REGION Network 31: Positioning commands
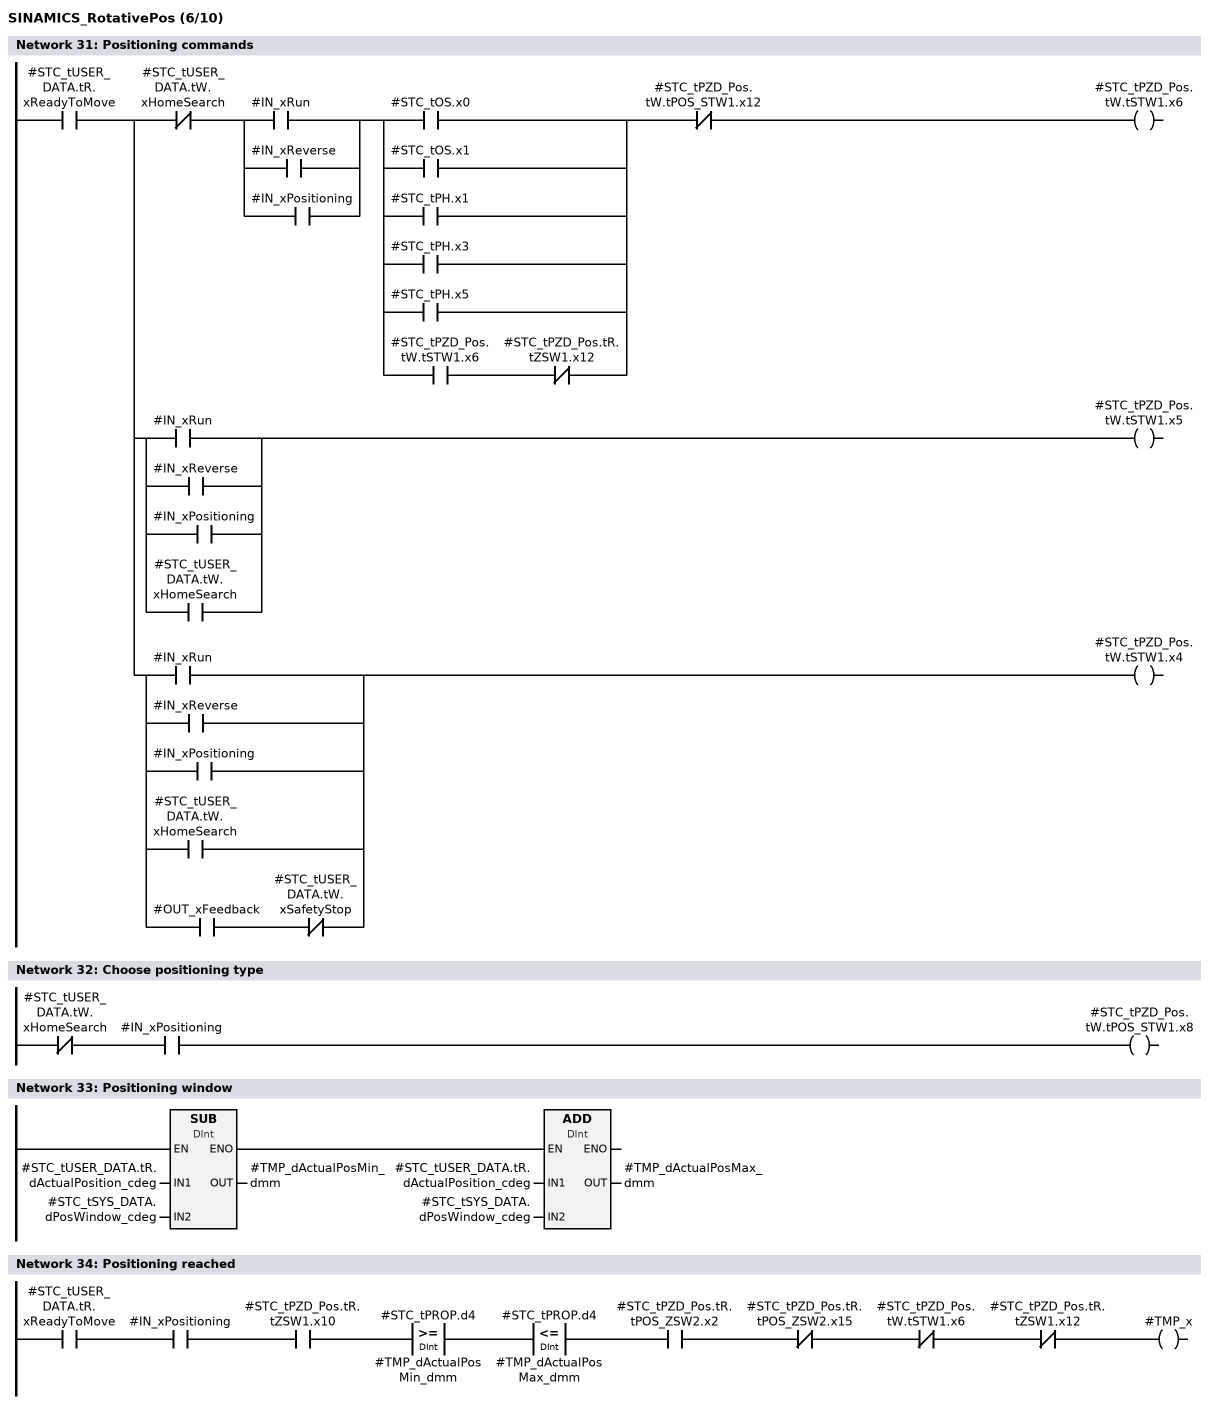
   RUNG wire#powerrail
      Contact( #STC_tUSER_DATA.tR.xReadyToMove )
      wire#w1
      I_Contact( #STC_tUSER_DATA.tW.xHomeSearch )
      wire#w2
      Contact( #IN_xRun )
      wire#w3
      Contact( #STC_tOS.x0 )
      wire#w4
      I_Contact( #STC_tPZD_Pos.tW.tPOS_STW1.x12 )
      Coil( #STC_tPZD_Pos.tW.tSTW1.x6 )
   END_RUNG
   RUNG wire#w2
      Contact( #IN_xReverse )
   END_RUNG wire#w3
   RUNG wire#w2
      Contact( #IN_xPositioning )
   END_RUNG wire#w3
   RUNG wire#w3
      Contact( #STC_tOS.x1 )
   END_RUNG wire#w4
   RUNG wire#w3
      Contact( #STC_tPH.x1 )
   END_RUNG wire#w4
   RUNG wire#w3
      Contact( #STC_tPH.x3 )
   END_RUNG wire#w4
   RUNG wire#w3
      Contact( #STC_tPH.x5 )
   END_RUNG wire#w4
   RUNG wire#w3
      Contact( #STC_tPZD_Pos.tW.tSTW1.x6 )
      I_Contact( #STC_tPZD_Pos.tR.tZSW1.x12 )
   END_RUNG wire#w4
   RUNG wire#w1
      Contact( #IN_xRun )
      wire#w5
      Coil( #STC_tPZD_Pos.tW.tSTW1.x5 )
   END_RUNG
   RUNG wire#w1
      Contact( #IN_xReverse )
   END_RUNG wire#w5
   RUNG wire#w1
      Contact( #IN_xPositioning )
   END_RUNG wire#w5
   RUNG wire#w1
      Contact( #STC_tUSER_DATA.tW.xHomeSearch )
   END_RUNG wire#w5
   RUNG wire#w1
      Contact( #IN_xRun )
      wire#w6
      Coil( #STC_tPZD_Pos.tW.tSTW1.x4 )
   END_RUNG
   RUNG wire#w1
      Contact( #IN_xReverse )
   END_RUNG wire#w6
   RUNG wire#w1
      Contact( #IN_xPositioning )
   END_RUNG wire#w6
   RUNG wire#w1
      Contact( #STC_tUSER_DATA.tW.xHomeSearch )
   END_RUNG wire#w6
   RUNG wire#w1
      Contact( #OUT_xFeedback )
      I_Contact( #STC_tUSER_DATA.tW.xSafetyStop )
   END_RUNG wire#w6
   // the same network as SCL:
   #STC_tPZD_Pos.tW.tSTW1.x6 := #STC_tUSER_DATA.tR.xReadyToMove AND NOT #STC_tUSER_DATA.tW.xHomeSearch AND (#IN_xRun OR #IN_xReverse OR #IN_xPositioning) AND (#STC_tOS.x0 OR #STC_tOS.x1 OR #STC_tPH.x1 OR #STC_tPH.x3 OR #STC_tPH.x5 OR (#STC_tPZD_Pos.tW.tSTW1.x6 AND NOT #STC_tPZD_Pos.tR.tZSW1.x12)) AND NOT #STC_tPZD_Pos.tW.tPOS_STW1.x12;
   #STC_tPZD_Pos.tW.tSTW1.x5 := #STC_tUSER_DATA.tR.xReadyToMove AND (#IN_xRun OR #IN_xReverse OR #IN_xPositioning OR #STC_tUSER_DATA.tW.xHomeSearch);
   #STC_tPZD_Pos.tW.tSTW1.x4 := #STC_tUSER_DATA.tR.xReadyToMove AND (#IN_xRun OR #IN_xReverse OR #IN_xPositioning OR #STC_tUSER_DATA.tW.xHomeSearch OR (#OUT_xFeedback AND NOT #STC_tUSER_DATA.tW.xSafetyStop));
END_REGION

REGION Network 32: Choose positioning type
   RUNG wire#powerrail
      I_Contact( #STC_tUSER_DATA.tW.xHomeSearch )
      Contact( #IN_xPositioning )
      Coil( #STC_tPZD_Pos.tW.tPOS_STW1.x8 )
   END_RUNG
   // the same network as SCL:
   #STC_tPZD_Pos.tW.tPOS_STW1.x8 := NOT #STC_tUSER_DATA.tW.xHomeSearch AND #IN_xPositioning;
END_REGION

REGION Network 33: Positioning window
   RUNG wire#powerrail
      { S7_Templates := "SrcType := DInt"; S7_GenerateENO := "TRUE" } Sub(in1 := #STC_tUSER_DATA.tR.dActualPosition_cdeg, in2 := #STC_tSYS_DATA.dPosWindow_cdeg, out => #TMP_dActualPosMin_dmm)
      { S7_Templates := "SrcType := DInt"; S7_GenerateENO := "TRUE" } Add(in1 := #STC_tUSER_DATA.tR.dActualPosition_cdeg, in2 := #STC_tSYS_DATA.dPosWindow_cdeg, out => #TMP_dActualPosMax_dmm)
   END_RUNG
   // the same network as SCL:
   // ENO of a box is taken as its EN; it also drops when the box reports an error
   #TMP_dActualPosMin_dmm := #STC_tUSER_DATA.tR.dActualPosition_cdeg - #STC_tSYS_DATA.dPosWindow_cdeg;
   #TMP_dActualPosMax_dmm := #STC_tUSER_DATA.tR.dActualPosition_cdeg + #STC_tSYS_DATA.dPosWindow_cdeg;
END_REGION

REGION Network 34: Positioning reached
   RUNG wire#powerrail
      Contact( #STC_tUSER_DATA.tR.xReadyToMove )
      Contact( #IN_xPositioning )
      Contact( #STC_tPZD_Pos.tR.tZSW1.x10 )
      { S7_Templates := "SrcType := DInt" } GE_Contact(in1 := #STC_tPROP.d4, in2 := #TMP_dActualPosMin_dmm)
      { S7_Templates := "SrcType := DInt" } LE_Contact(in1 := #STC_tPROP.d4, in2 := #TMP_dActualPosMax_dmm)
      Contact( #STC_tPZD_Pos.tR.tPOS_ZSW2.x2 )
      I_Contact( #STC_tPZD_Pos.tR.tPOS_ZSW2.x15 )
      I_Contact( #STC_tPZD_Pos.tW.tSTW1.x6 )
      I_Contact( #STC_tPZD_Pos.tR.tZSW1.x12 )
      Coil( #TMP_x )
   END_RUNG
   // the same network as SCL:
   #TMP_x := #STC_tUSER_DATA.tR.xReadyToMove AND #IN_xPositioning AND #STC_tPZD_Pos.tR.tZSW1.x10 AND (#STC_tPROP.d4 >= #TMP_dActualPosMin_dmm) AND (#STC_tPROP.d4 <= #TMP_dActualPosMax_dmm) AND #STC_tPZD_Pos.tR.tPOS_ZSW2.x2 AND NOT #STC_tPZD_Pos.tR.tPOS_ZSW2.x15 AND NOT #STC_tPZD_Pos.tW.tSTW1.x6 AND NOT #STC_tPZD_Pos.tR.tZSW1.x12;
END_REGION

REGION Network 35: Positioning reached
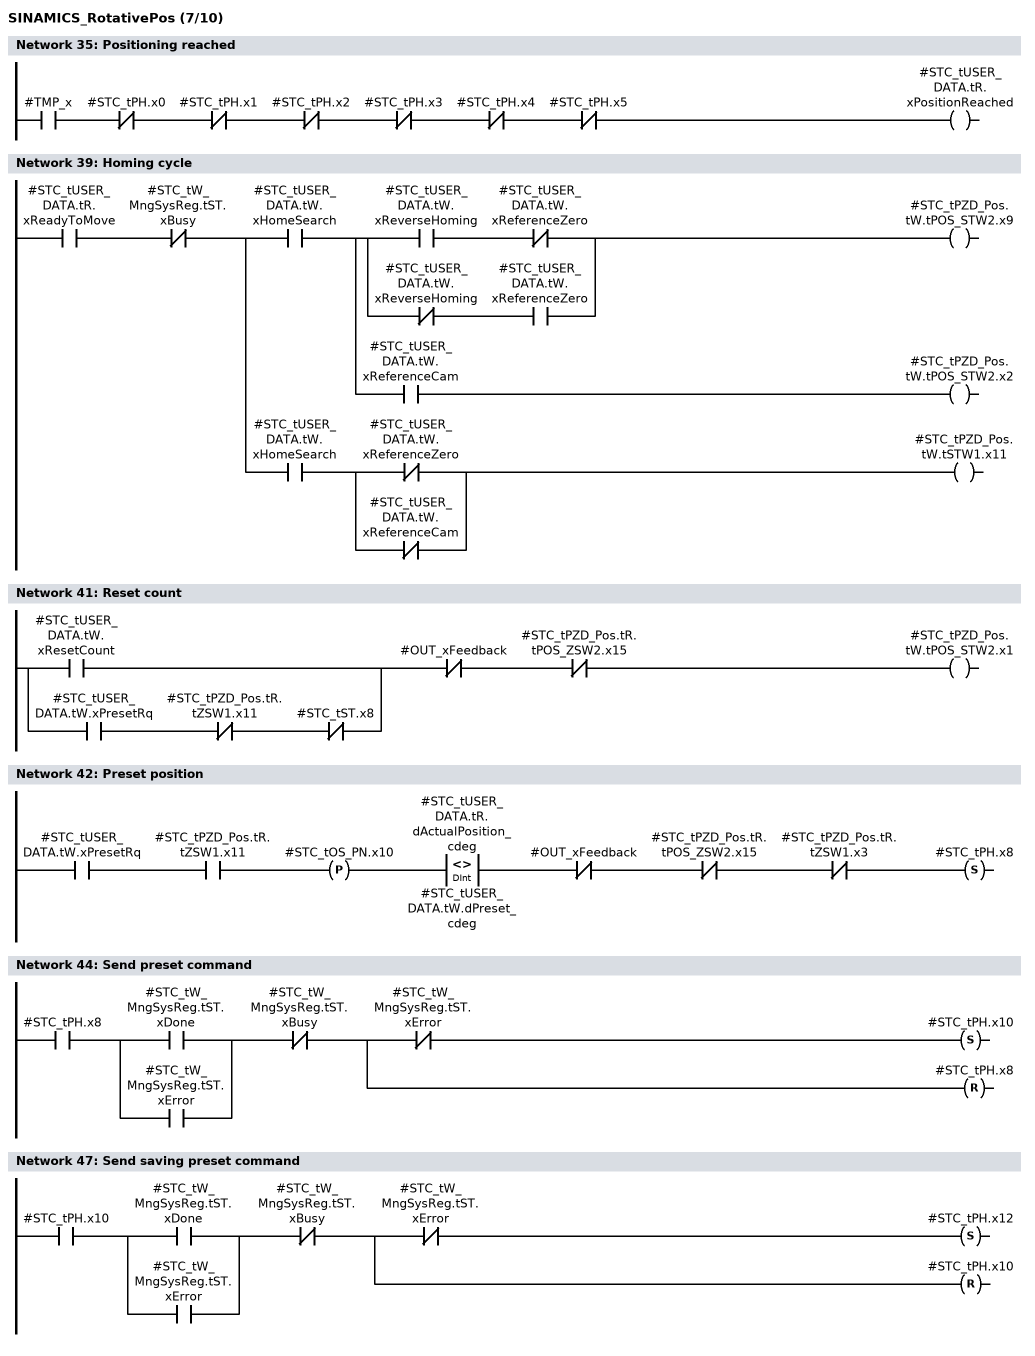
   RUNG wire#powerrail
      Contact( #TMP_x )
      I_Contact( #STC_tPH.x0 )
      I_Contact( #STC_tPH.x1 )
      I_Contact( #STC_tPH.x2 )
      I_Contact( #STC_tPH.x3 )
      I_Contact( #STC_tPH.x4 )
      I_Contact( #STC_tPH.x5 )
      Coil( #STC_tUSER_DATA.tR.xPositionReached )
   END_RUNG
   // the same network as SCL:
   #STC_tUSER_DATA.tR.xPositionReached := #TMP_x AND NOT #STC_tPH.x0 AND NOT #STC_tPH.x1 AND NOT #STC_tPH.x2 AND NOT #STC_tPH.x3 AND NOT #STC_tPH.x4 AND NOT #STC_tPH.x5;
END_REGION

REGION Network 36: #####_HOMING_CYCLE_#####
END_REGION

REGION Network 37 (STL): Send homing preset
         A     #STC_tUSER_DATA.tW.xHomeSearch;
         AN    #STC_tPZD_Pos.tW.tSTW1.x11;
         JCN   PrH0;
         =     #STC_tW_MngSysReg.tST.xWrite_Request;

         L     #STC_tSYS_DATA.iPosPZD_MM;
         SLW   8;
         L     W#16#2;
         OW;
         T     #STC_tW_MngSysReg.tDATA.wRequest_refere_RequestID;
         L     #STC_tSYS_DATA.iPosPZD_MM;
         SLW   8;
         L     W#16#1;
         OW;
         T     #STC_tW_MngSysReg.tDATA.wAxis_NoOfParameters;
         L     W#16#1001;
         T     #STC_tW_MngSysReg.tDATA.wAttribute_NoOfElements;
         L     2599;
         T     #STC_tW_MngSysReg.tDATA.iParameter_number;
         L     W#16#0;
         T     #STC_tW_MngSysReg.tDATA.wSubindex;
         L     W#16#4301;
         T     #STC_tW_MngSysReg.tDATA.wFormat_NoOfValue;
         L     #STC_tSYS_DATA.iDiagAddress;
         T     #STC_tW_MngSysReg.tST.ID;
         L     47;
         T     #STC_tW_MngSysReg.tST.dINDEX;
         L     16;
         T     #STC_tW_MngSysReg.tST.uiLEN;

         L     #STC_tUSER_DATA.tW.dPreset_cdeg;
         T     #STC_tW_MngSysReg.tDATA.dwRegisterValue;

         CALL  #STC_tWriteRecord
         ( REQ    := #STC_tW_MngSysReg.tST.xWrite_Request,
           ID     := #STC_tW_MngSysReg.tST.ID,
           INDEX  := #STC_tW_MngSysReg.tST.dINDEX,
           LEN    := #STC_tW_MngSysReg.tST.uiLEN,
           DONE   := #STC_tW_MngSysReg.tST.xDone,
           BUSY   := #STC_tW_MngSysReg.tST.xBusy,
           ERROR  := #STC_tW_MngSysReg.tST.xError,
           STATUS := #STC_tW_MngSysReg.tST.dwSTATUS,
           RECORD := #STC_tW_MngSysReg.tDATA
         );
   PrH0: NOP   0;
END_REGION

REGION Network 38 (STL): Error during Send homing preset
         A     #STC_tW_MngSysReg.tST.xError;
         L     34;
         JC    Err;
END_REGION

REGION Network 39: Homing cycle
   RUNG wire#powerrail
      Contact( #STC_tUSER_DATA.tR.xReadyToMove )
      I_Contact( #STC_tW_MngSysReg.tST.xBusy )
      wire#w1
      Contact( #STC_tUSER_DATA.tW.xHomeSearch )
      wire#w2
      Contact( #STC_tUSER_DATA.tW.xReverseHoming )
      I_Contact( #STC_tUSER_DATA.tW.xReferenceZero )
      wire#w3
      Coil( #STC_tPZD_Pos.tW.tPOS_STW2.x9 )
   END_RUNG
   RUNG wire#w2
      I_Contact( #STC_tUSER_DATA.tW.xReverseHoming )
      Contact( #STC_tUSER_DATA.tW.xReferenceZero )
   END_RUNG wire#w3
   RUNG wire#w2
      Contact( #STC_tUSER_DATA.tW.xReferenceCam )
      Coil( #STC_tPZD_Pos.tW.tPOS_STW2.x2 )
   END_RUNG
   RUNG wire#w1
      Contact( #STC_tUSER_DATA.tW.xHomeSearch )
      wire#w4
      I_Contact( #STC_tUSER_DATA.tW.xReferenceZero )
      wire#w5
      Coil( #STC_tPZD_Pos.tW.tSTW1.x11 )
   END_RUNG
   RUNG wire#w4
      I_Contact( #STC_tUSER_DATA.tW.xReferenceCam )
   END_RUNG wire#w5
   // the same network as SCL:
   #_w1 := #STC_tUSER_DATA.tR.xReadyToMove AND NOT #STC_tW_MngSysReg.tST.xBusy;
   #_w2 := #_w1 AND #STC_tUSER_DATA.tW.xHomeSearch;
   #STC_tPZD_Pos.tW.tPOS_STW2.x9 := #_w2 AND ((#STC_tUSER_DATA.tW.xReverseHoming AND NOT #STC_tUSER_DATA.tW.xReferenceZero) OR (NOT #STC_tUSER_DATA.tW.xReverseHoming AND #STC_tUSER_DATA.tW.xReferenceZero));
   #STC_tPZD_Pos.tW.tPOS_STW2.x2 := #_w2 AND #STC_tUSER_DATA.tW.xReferenceCam;
   #STC_tPZD_Pos.tW.tSTW1.x11 := #_w1 AND #STC_tUSER_DATA.tW.xHomeSearch AND (NOT #STC_tUSER_DATA.tW.xReferenceZero OR NOT #STC_tUSER_DATA.tW.xReferenceCam);
END_REGION

REGION Network 40: #####_PRESET_ACTUAL_POSITION_#####
END_REGION

REGION Network 41: Reset count
   RUNG wire#powerrail
      Contact( #STC_tUSER_DATA.tW.xResetCount )
      wire#w1
      I_Contact( #OUT_xFeedback )
      I_Contact( #STC_tPZD_Pos.tR.tPOS_ZSW2.x15 )
      Coil( #STC_tPZD_Pos.tW.tPOS_STW2.x1 )
   END_RUNG
   RUNG wire#powerrail
      Contact( #STC_tUSER_DATA.tW.xPresetRq )
      I_Contact( #STC_tPZD_Pos.tR.tZSW1.x11 )
      I_Contact( #STC_tST.x8 )
   END_RUNG wire#w1
   // the same network as SCL:
   #STC_tPZD_Pos.tW.tPOS_STW2.x1 := (#STC_tUSER_DATA.tW.xResetCount OR (#STC_tUSER_DATA.tW.xPresetRq AND NOT #STC_tPZD_Pos.tR.tZSW1.x11 AND NOT #STC_tST.x8)) AND NOT #OUT_xFeedback AND NOT #STC_tPZD_Pos.tR.tPOS_ZSW2.x15;
END_REGION

REGION Network 42: Preset position
   RUNG wire#powerrail
      Contact( #STC_tUSER_DATA.tW.xPresetRq )
      Contact( #STC_tPZD_Pos.tR.tZSW1.x11 )
      P_Trig( #STC_tOS_PN.x10 )
      { S7_Templates := "SrcType := DInt" } NE_Contact(in1 := #STC_tUSER_DATA.tR.dActualPosition_cdeg, in2 := #STC_tUSER_DATA.tW.dPreset_cdeg)
      I_Contact( #OUT_xFeedback )
      I_Contact( #STC_tPZD_Pos.tR.tPOS_ZSW2.x15 )
      I_Contact( #STC_tPZD_Pos.tR.tZSW1.x3 )
      S_Coil( #STC_tPH.x8 )
   END_RUNG
   // the same network as SCL:
   #_w1 := #STC_tUSER_DATA.tW.xPresetRq AND #STC_tPZD_Pos.tR.tZSW1.x11;
   #_w2 := #_w1 AND NOT #STC_tOS_PN.x10;   // rising edge
   #STC_tOS_PN.x10 := #_w1;
   IF #_w2 AND (#STC_tUSER_DATA.tR.dActualPosition_cdeg <> #STC_tUSER_DATA.tW.dPreset_cdeg) AND NOT #OUT_xFeedback AND NOT #STC_tPZD_Pos.tR.tPOS_ZSW2.x15 AND NOT #STC_tPZD_Pos.tR.tZSW1.x3 THEN
       #STC_tPH.x8 := TRUE;
   END_IF;
END_REGION

REGION Network 43 (STL): Send encoder value
         A     #STC_tPH.x8;
         JCN   PrE0;
         =     #STC_tW_MngSysReg.tST.xWrite_Request;

         L     #STC_tSYS_DATA.iPosPZD_MM;
         +     10;
         SLW   8;
         L     W#16#2;
         OW;
         T     #STC_tW_MngSysReg.tDATA.wRequest_refere_RequestID;
         L     #STC_tSYS_DATA.iPosPZD_MM;
         SLW   8;
         L     W#16#1;
         OW;
         T     #STC_tW_MngSysReg.tDATA.wAxis_NoOfParameters;
         L     W#16#1001;
         T     #STC_tW_MngSysReg.tDATA.wAttribute_NoOfElements;
         L     2599;
         T     #STC_tW_MngSysReg.tDATA.iParameter_number;
         L     W#16#0;
         T     #STC_tW_MngSysReg.tDATA.wSubindex;
         L     W#16#4301;
         T     #STC_tW_MngSysReg.tDATA.wFormat_NoOfValue;
         L     #STC_tSYS_DATA.iDiagAddress;
         T     #STC_tW_MngSysReg.tST.ID;
         L     47;
         T     #STC_tW_MngSysReg.tST.dINDEX;
         L     16;
         T     #STC_tW_MngSysReg.tST.uiLEN;

         L     #STC_tUSER_DATA.tW.dPreset_cdeg;
         T     #STC_tW_MngSysReg.tDATA.dwRegisterValue;

         CALL  #STC_tWriteRecord
         ( REQ    := #STC_tW_MngSysReg.tST.xWrite_Request,
           ID     := #STC_tW_MngSysReg.tST.ID,
           INDEX  := #STC_tW_MngSysReg.tST.dINDEX,
           LEN    := #STC_tW_MngSysReg.tST.uiLEN,
           DONE   := #STC_tW_MngSysReg.tST.xDone,
           BUSY   := #STC_tW_MngSysReg.tST.xBusy,
           ERROR  := #STC_tW_MngSysReg.tST.xError,
           STATUS := #STC_tW_MngSysReg.tST.dwSTATUS,
           RECORD := #STC_tW_MngSysReg.tDATA
         );
   PrE0: NOP   0;
END_REGION

REGION Network 44: Send preset command
   RUNG wire#powerrail
      Contact( #STC_tPH.x8 )
      wire#w1
      Contact( #STC_tW_MngSysReg.tST.xDone )
      wire#w2
      I_Contact( #STC_tW_MngSysReg.tST.xBusy )
      wire#w3
      I_Contact( #STC_tW_MngSysReg.tST.xError )
      S_Coil( #STC_tPH.x10 )
   END_RUNG
   RUNG wire#w1
      Contact( #STC_tW_MngSysReg.tST.xError )
   END_RUNG wire#w2
   RUNG wire#w3
      R_Coil( #STC_tPH.x8 )
   END_RUNG
   // the same network as SCL:
   #_w1 := #STC_tPH.x8 AND (#STC_tW_MngSysReg.tST.xDone OR #STC_tW_MngSysReg.tST.xError) AND NOT #STC_tW_MngSysReg.tST.xBusy;
   IF #_w1 AND NOT #STC_tW_MngSysReg.tST.xError THEN #STC_tPH.x10 := TRUE; END_IF;
   IF #_w1 THEN #STC_tPH.x8 := FALSE; END_IF;
END_REGION

REGION Network 45 (STL): Error during send ecoder value
         A     #STC_tW_MngSysReg.tST.xError;
         L     30;
         JC    Err;
END_REGION

REGION Network 46 (STL): Send preset command
         A     #STC_tPH.x10;
         JCN   PrE1;
         =     #STC_tW_MngSysReg.tST.xWrite_Request;

         L     #STC_tSYS_DATA.iPosPZD_MM;
         +     20;
         SLW   8;
         L     W#16#2;
         OW;
         T     #STC_tW_MngSysReg.tDATA.wRequest_refere_RequestID;
         L     #STC_tSYS_DATA.iPosPZD_MM;
         SLW   8;
         L     W#16#1;
         OW;
         T     #STC_tW_MngSysReg.tDATA.wAxis_NoOfParameters;
         L     W#16#1001;
         T     #STC_tW_MngSysReg.tDATA.wAttribute_NoOfElements;
         L     2507;
         T     #STC_tW_MngSysReg.tDATA.iParameter_number;
         L     W#16#0;
         T     #STC_tW_MngSysReg.tDATA.wSubindex;
         L     W#16#4201;
         T     #STC_tW_MngSysReg.tDATA.wFormat_NoOfValue;
         L     #STC_tSYS_DATA.iDiagAddress;
         T     #STC_tW_MngSysReg.tST.ID;
         L     47;
         T     #STC_tW_MngSysReg.tST.dINDEX;
         L     14;
         T     #STC_tW_MngSysReg.tST.uiLEN;

         L     DINT#2;
         SLD   16;
         T     #STC_tW_MngSysReg.tDATA.dwRegisterValue;

         CALL  #STC_tWriteRecord
         ( REQ    := #STC_tW_MngSysReg.tST.xWrite_Request,
           ID     := #STC_tW_MngSysReg.tST.ID,
           INDEX  := #STC_tW_MngSysReg.tST.dINDEX,
           LEN    := #STC_tW_MngSysReg.tST.uiLEN,
           DONE   := #STC_tW_MngSysReg.tST.xDone,
           BUSY   := #STC_tW_MngSysReg.tST.xBusy,
           ERROR  := #STC_tW_MngSysReg.tST.xError,
           STATUS := #STC_tW_MngSysReg.tST.dwSTATUS,
           RECORD := #STC_tW_MngSysReg.tDATA
         );
   PrE1: NOP   0;
END_REGION

REGION Network 47: Send saving preset command
   RUNG wire#powerrail
      Contact( #STC_tPH.x10 )
      wire#w1
      Contact( #STC_tW_MngSysReg.tST.xDone )
      wire#w2
      I_Contact( #STC_tW_MngSysReg.tST.xBusy )
      wire#w3
      I_Contact( #STC_tW_MngSysReg.tST.xError )
      S_Coil( #STC_tPH.x12 )
   END_RUNG
   RUNG wire#w1
      Contact( #STC_tW_MngSysReg.tST.xError )
   END_RUNG wire#w2
   RUNG wire#w3
      R_Coil( #STC_tPH.x10 )
   END_RUNG
   // the same network as SCL:
   #_w1 := #STC_tPH.x10 AND (#STC_tW_MngSysReg.tST.xDone OR #STC_tW_MngSysReg.tST.xError) AND NOT #STC_tW_MngSysReg.tST.xBusy;
   IF #_w1 AND NOT #STC_tW_MngSysReg.tST.xError THEN #STC_tPH.x12 := TRUE; END_IF;
   IF #_w1 THEN #STC_tPH.x10 := FALSE; END_IF;
END_REGION

REGION Network 48 (STL): Error during preset command
         A     #STC_tW_MngSysReg.tST.xError;
         L     31;
         JC    Err;
END_REGION

REGION Network 49 (STL): Send saving preset command
         A     #STC_tPH.x12;
         JCN   PrE2;
         =     #STC_tW_MngSysReg.tST.xWrite_Request;

         L     #STC_tSYS_DATA.iPosPZD_MM;
         +     30;
         SLW   8;
         L     W#16#2;
         OW;
         T     #STC_tW_MngSysReg.tDATA.wRequest_refere_RequestID;
         L     #STC_tSYS_DATA.iPosPZD_CU;
         SLW   8;
         L     W#16#1;
         OW;
         T     #STC_tW_MngSysReg.tDATA.wAxis_NoOfParameters;
         L     W#16#1001;
         T     #STC_tW_MngSysReg.tDATA.wAttribute_NoOfElements;
         L     977;
         T     #STC_tW_MngSysReg.tDATA.iParameter_number;
         L     W#16#0;
         T     #STC_tW_MngSysReg.tDATA.wSubindex;
         L     W#16#4201;
         T     #STC_tW_MngSysReg.tDATA.wFormat_NoOfValue;
         L     #STC_tSYS_DATA.iDiagAddress;
         T     #STC_tW_MngSysReg.tST.ID;
         L     47;
         T     #STC_tW_MngSysReg.tST.dINDEX;
         L     14;
         T     #STC_tW_MngSysReg.tST.uiLEN;

         L     DINT#1;
         SLD   16;
         T     #STC_tW_MngSysReg.tDATA.dwRegisterValue;

         CALL  #STC_tWriteRecord
         ( REQ    := #STC_tW_MngSysReg.tST.xWrite_Request,
           ID     := #STC_tW_MngSysReg.tST.ID,
           INDEX  := #STC_tW_MngSysReg.tST.dINDEX,
           LEN    := #STC_tW_MngSysReg.tST.uiLEN,
           DONE   := #STC_tW_MngSysReg.tST.xDone,
           BUSY   := #STC_tW_MngSysReg.tST.xBusy,
           ERROR  := #STC_tW_MngSysReg.tST.xError,
           STATUS := #STC_tW_MngSysReg.tST.dwSTATUS,
           RECORD := #STC_tW_MngSysReg.tDATA
         );
   PrE2: NOP   0;
END_REGION

REGION Network 50: End preset encoder
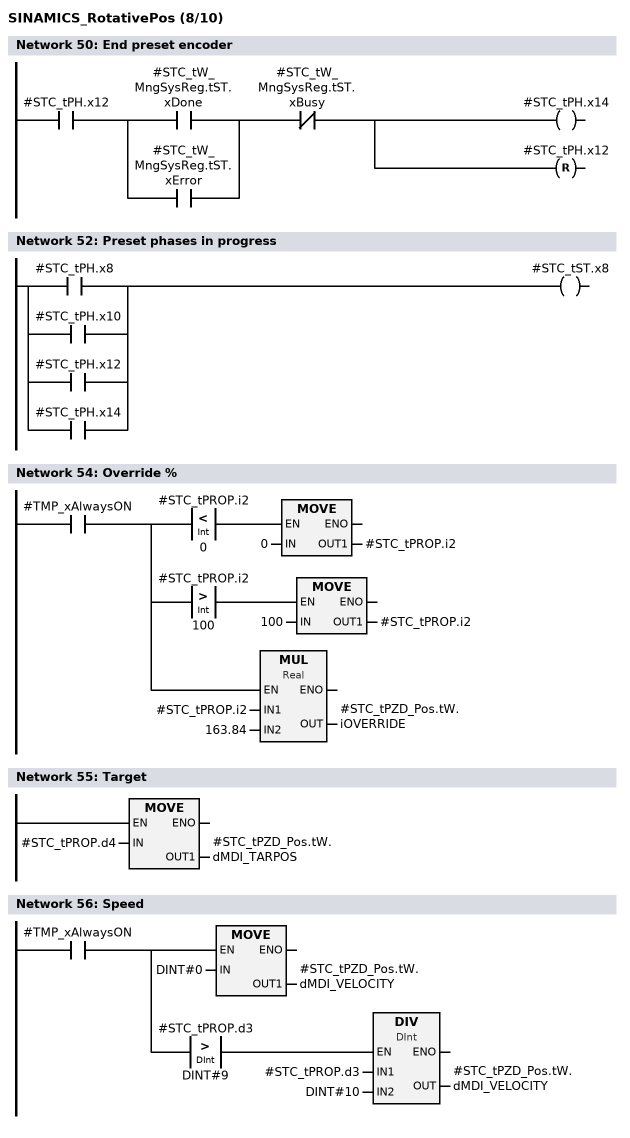
   RUNG wire#powerrail
      Contact( #STC_tPH.x12 )
      wire#w1
      Contact( #STC_tW_MngSysReg.tST.xDone )
      wire#w2
      I_Contact( #STC_tW_MngSysReg.tST.xBusy )
      wire#w3
      Coil( #STC_tPH.x14 )
   END_RUNG
   RUNG wire#w1
      Contact( #STC_tW_MngSysReg.tST.xError )
   END_RUNG wire#w2
   RUNG wire#w3
      R_Coil( #STC_tPH.x12 )
   END_RUNG
   // the same network as SCL:
   #STC_tPH.x14 := #STC_tPH.x12 AND (#STC_tW_MngSysReg.tST.xDone OR #STC_tW_MngSysReg.tST.xError) AND NOT #STC_tW_MngSysReg.tST.xBusy;
   IF #STC_tPH.x14 THEN #STC_tPH.x12 := FALSE; END_IF;
END_REGION

REGION Network 51 (STL): Error during saving preset command
         A     #STC_tW_MngSysReg.tST.xError;
         L     32;
         JC    Err;
END_REGION

REGION Network 52: Preset phases in progress
   RUNG wire#powerrail
      Contact( #STC_tPH.x8 )
      wire#w1
      Coil( #STC_tST.x8 )
   END_RUNG
   RUNG wire#powerrail
      Contact( #STC_tPH.x10 )
   END_RUNG wire#w1
   RUNG wire#powerrail
      Contact( #STC_tPH.x12 )
   END_RUNG wire#w1
   RUNG wire#powerrail
      Contact( #STC_tPH.x14 )
   END_RUNG wire#w1
   // the same network as SCL:
   #STC_tST.x8 := #STC_tPH.x8 OR #STC_tPH.x10 OR #STC_tPH.x12 OR #STC_tPH.x14;
END_REGION

REGION Network 53: #####_PARAMETERS_#####
END_REGION

REGION Network 54: Override %
   RUNG wire#powerrail
      Contact( #TMP_xAlwaysON )
      wire#w1
      { S7_Templates := "SrcType := Int" } LT_Contact(in1 := #STC_tPROP.i2, in2 := 0)
      Move(in := 0, out1 => #STC_tPROP.i2)
   END_RUNG
   RUNG wire#w1
      { S7_Templates := "SrcType := Int" } GT_Contact(in1 := #STC_tPROP.i2, in2 := 100)
      Move(in := 100, out1 => #STC_tPROP.i2)
   END_RUNG
   RUNG wire#w1
      { S7_Templates := "SrcType := Real" } Mul(in1 := #STC_tPROP.i2, in2 := 163.84, out => #STC_tPZD_Pos.tW.iOVERRIDE)
   END_RUNG
   // the same network as SCL:
   IF #TMP_xAlwaysON AND (#STC_tPROP.i2 < 0) THEN #STC_tPROP.i2 := 0; END_IF;
   IF #TMP_xAlwaysON AND (#STC_tPROP.i2 > 100) THEN #STC_tPROP.i2 := 100; END_IF;
   IF #TMP_xAlwaysON THEN #STC_tPZD_Pos.tW.iOVERRIDE := #STC_tPROP.i2 * 163.84; END_IF;
END_REGION

REGION Network 55: Target
   RUNG wire#powerrail
      { S7_GenerateENO := "TRUE" } Move(in := #STC_tPROP.d4, out1 => #STC_tPZD_Pos.tW.dMDI_TARPOS)
   END_RUNG
   // the same network as SCL:
   #STC_tPZD_Pos.tW.dMDI_TARPOS := #STC_tPROP.d4;
END_REGION

REGION Network 56: Speed
   RUNG wire#powerrail
      Contact( #TMP_xAlwaysON )
      wire#w1
      { S7_GenerateENO := "TRUE" } Move(in := DINT#0, out1 => #STC_tPZD_Pos.tW.dMDI_VELOCITY)
   END_RUNG
   RUNG wire#w1
      { S7_Templates := "SrcType := DInt" } GT_Contact(in1 := #STC_tPROP.d3, in2 := DINT#9)
      { S7_Templates := "SrcType := DInt"; S7_GenerateENO := "TRUE" } Div(in1 := #STC_tPROP.d3, in2 := DINT#10, out => #STC_tPZD_Pos.tW.dMDI_VELOCITY)
   END_RUNG
   // the same network as SCL:
   IF #TMP_xAlwaysON THEN #STC_tPZD_Pos.tW.dMDI_VELOCITY := DINT#0; END_IF;
   IF #TMP_xAlwaysON AND (#STC_tPROP.d3 > DINT#9) THEN
       #STC_tPZD_Pos.tW.dMDI_VELOCITY := #STC_tPROP.d3 / DINT#10;
   END_IF;
END_REGION

REGION Network 57: Acceleration
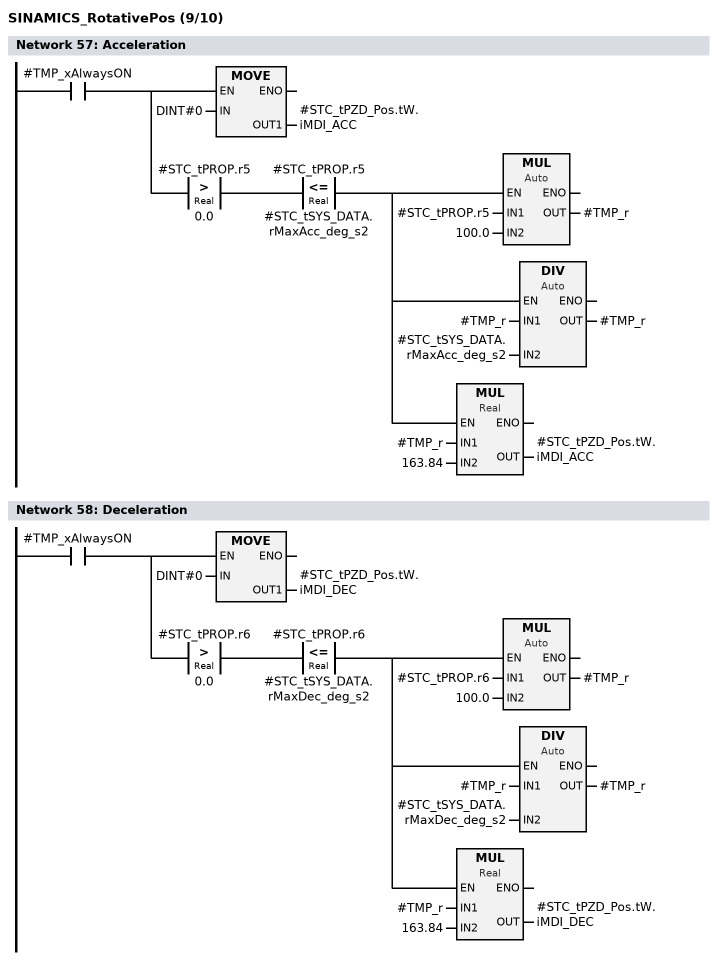
   RUNG wire#powerrail
      Contact( #TMP_xAlwaysON )
      wire#w1
      Move(in := DINT#0, out1 => #STC_tPZD_Pos.tW.iMDI_ACC)
   END_RUNG
   RUNG wire#w1
      { S7_Templates := "SrcType := Real" } GT_Contact(in1 := #STC_tPROP.r5, in2 := 0.0)
      { S7_Templates := "SrcType := Real" } LE_Contact(in1 := #STC_tPROP.r5, in2 := #STC_tSYS_DATA.rMaxAcc_deg_s2)
      wire#w2
      Mul(in1 := #STC_tPROP.r5, in2 := 100.0, out => #TMP_r)
   END_RUNG
   RUNG wire#w2
      Div(in1 := #TMP_r, in2 := #STC_tSYS_DATA.rMaxAcc_deg_s2, out => #TMP_r)
   END_RUNG
   RUNG wire#w2
      { S7_Templates := "SrcType := Real" } Mul(in1 := #TMP_r, in2 := 163.84, out => #STC_tPZD_Pos.tW.iMDI_ACC)
   END_RUNG
   // the same network as SCL:
   IF #TMP_xAlwaysON THEN #STC_tPZD_Pos.tW.iMDI_ACC := DINT#0; END_IF;
   IF #TMP_xAlwaysON AND (#STC_tPROP.r5 > 0.0) AND (#STC_tPROP.r5 <= #STC_tSYS_DATA.rMaxAcc_deg_s2) THEN
       #TMP_r := #STC_tPROP.r5 * 100.0;
       #TMP_r := #TMP_r / #STC_tSYS_DATA.rMaxAcc_deg_s2;
       #STC_tPZD_Pos.tW.iMDI_ACC := #TMP_r * 163.84;
   END_IF;
END_REGION

REGION Network 58: Deceleration
   RUNG wire#powerrail
      Contact( #TMP_xAlwaysON )
      wire#w1
      Move(in := DINT#0, out1 => #STC_tPZD_Pos.tW.iMDI_DEC)
   END_RUNG
   RUNG wire#w1
      { S7_Templates := "SrcType := Real" } GT_Contact(in1 := #STC_tPROP.r6, in2 := 0.0)
      { S7_Templates := "SrcType := Real" } LE_Contact(in1 := #STC_tPROP.r6, in2 := #STC_tSYS_DATA.rMaxDec_deg_s2)
      wire#w2
      Mul(in1 := #STC_tPROP.r6, in2 := 100.0, out => #TMP_r)
   END_RUNG
   RUNG wire#w2
      Div(in1 := #TMP_r, in2 := #STC_tSYS_DATA.rMaxDec_deg_s2, out => #TMP_r)
   END_RUNG
   RUNG wire#w2
      { S7_Templates := "SrcType := Real" } Mul(in1 := #TMP_r, in2 := 163.84, out => #STC_tPZD_Pos.tW.iMDI_DEC)
   END_RUNG
   // the same network as SCL:
   IF #TMP_xAlwaysON THEN #STC_tPZD_Pos.tW.iMDI_DEC := DINT#0; END_IF;
   IF #TMP_xAlwaysON AND (#STC_tPROP.r6 > 0.0) AND (#STC_tPROP.r6 <= #STC_tSYS_DATA.rMaxDec_deg_s2) THEN
       #TMP_r := #STC_tPROP.r6 * 100.0;
       #TMP_r := #TMP_r / #STC_tSYS_DATA.rMaxDec_deg_s2;
       #STC_tPZD_Pos.tW.iMDI_DEC := #TMP_r * 163.84;
   END_IF;
END_REGION

REGION Network 59: ################_MOTOR_MODULE_TELEGRAMS_ENDING_#################
END_REGION

REGION Network 60 (STL): Output copy motor module
   // Compute destination position
         L;
         LAR1;
   //byte 1 = 10h (FIXED for S7)
         L     B#16#10;
         T     B[AR1, P#0.0];
   //byte 2 = data type
         L     B#16#4;  //4 = word
         T     B[AR1, P#1.0];
   //byte 3 & 4 = number of element
         L     12;  //Production data
         T     W[AR1, P#2.0];
   //byte 5 & 6 = number of DB
         L     0;  //DB production data
         T     W[AR1, P#4.0];
   //byte 7 = memory area
         L     B#16#82;  //82h = Q (Output)
         T     B[AR1, P#6.0];
   //byte 8 & 9 = address. Bit 0,1,2 of tenth byte is bit offset
   //byte 7 = address (high). Valid value = 0-7. Bit 3,4,5,6,7 always 0
         L     #STC_tSYS_DATA.iIOAddress_MM;  //Item size
         SLW   3;
         T     W[AR1, P#8.0];
         SRD   16;
         AW    16#0007;
         T     B[AR1, P#7.0];

         CALL  BLKMOV
         ( SRCBLK  := #STC_tPZD_Pos.tW,
           RET_VAL := #TMP_iRetVal,
           DSTBLK  := #TMP_a
         );
END_REGION

REGION Network 61: #####_RETVAL_RESPONSE_#####
END_REGION

REGION Network 62 (STL): Initialize RetVal
         L     0;
         T     #OUT_iRetVal;
END_REGION

REGION Network 63: Warning messages
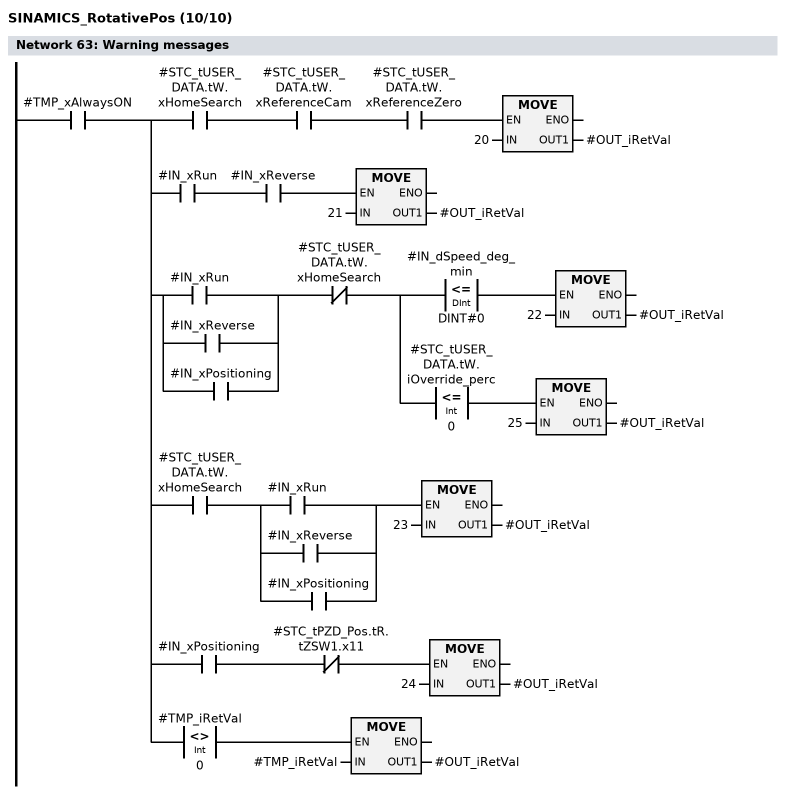
   RUNG wire#powerrail
      Contact( #TMP_xAlwaysON )
      wire#w1
      Contact( #STC_tUSER_DATA.tW.xHomeSearch )
      Contact( #STC_tUSER_DATA.tW.xReferenceCam )
      Contact( #STC_tUSER_DATA.tW.xReferenceZero )
      Move(in := 20, out1 => #OUT_iRetVal)
   END_RUNG
   RUNG wire#w1
      Contact( #IN_xRun )
      Contact( #IN_xReverse )
      Move(in := 21, out1 => #OUT_iRetVal)
   END_RUNG
   RUNG wire#w1
      Contact( #IN_xRun )
      wire#w2
      I_Contact( #STC_tUSER_DATA.tW.xHomeSearch )
      wire#w3
      { S7_Templates := "SrcType := DInt" } LE_Contact(in1 := #IN_dSpeed_deg_min, in2 := DINT#0)
      Move(in := 22, out1 => #OUT_iRetVal)
   END_RUNG
   RUNG wire#w1
      Contact( #IN_xReverse )
   END_RUNG wire#w2
   RUNG wire#w1
      Contact( #IN_xPositioning )
   END_RUNG wire#w2
   RUNG wire#w3
      { S7_Templates := "SrcType := Int" } LE_Contact(in1 := #STC_tUSER_DATA.tW.iOverride_perc, in2 := 0)
      Move(in := 25, out1 => #OUT_iRetVal)
   END_RUNG
   RUNG wire#w1
      Contact( #STC_tUSER_DATA.tW.xHomeSearch )
      wire#w4
      Contact( #IN_xRun )
      wire#w5
      Move(in := 23, out1 => #OUT_iRetVal)
   END_RUNG
   RUNG wire#w4
      Contact( #IN_xReverse )
   END_RUNG wire#w5
   RUNG wire#w4
      Contact( #IN_xPositioning )
   END_RUNG wire#w5
   RUNG wire#w1
      Contact( #IN_xPositioning )
      I_Contact( #STC_tPZD_Pos.tR.tZSW1.x11 )
      Move(in := 24, out1 => #OUT_iRetVal)
   END_RUNG
   RUNG wire#w1
      { S7_Templates := "SrcType := Int" } NE_Contact(in1 := #TMP_iRetVal, in2 := 0)
      Move(in := #TMP_iRetVal, out1 => #OUT_iRetVal)
   END_RUNG
   // the same network as SCL:
   IF #TMP_xAlwaysON AND #STC_tUSER_DATA.tW.xHomeSearch AND #STC_tUSER_DATA.tW.xReferenceCam AND #STC_tUSER_DATA.tW.xReferenceZero THEN
       #OUT_iRetVal := 20;
   END_IF;
   IF #TMP_xAlwaysON AND #IN_xRun AND #IN_xReverse THEN #OUT_iRetVal := 21; END_IF;
   #_w1 := #TMP_xAlwaysON AND (#IN_xRun OR #IN_xReverse OR #IN_xPositioning) AND NOT #STC_tUSER_DATA.tW.xHomeSearch;
   IF #_w1 AND (#IN_dSpeed_deg_min <= DINT#0) THEN #OUT_iRetVal := 22; END_IF;
   IF #_w1 AND (#STC_tUSER_DATA.tW.iOverride_perc <= 0) THEN #OUT_iRetVal := 25; END_IF;
   IF #TMP_xAlwaysON AND #STC_tUSER_DATA.tW.xHomeSearch AND (#IN_xRun OR #IN_xReverse OR #IN_xPositioning) THEN
       #OUT_iRetVal := 23;
   END_IF;
   IF #TMP_xAlwaysON AND #IN_xPositioning AND NOT #STC_tPZD_Pos.tR.tZSW1.x11 THEN #OUT_iRetVal := 24; END_IF;
   IF #TMP_xAlwaysON AND (#TMP_iRetVal <> 0) THEN #OUT_iRetVal := #TMP_iRetVal; END_IF;
END_REGION

REGION Network 64 (STL): Blocking messages
         JU    Rest;
   Err:  T     #OUT_iRetVal;
END_REGION

REGION Network 65 (STL): Reset input commands
   // R     #USER_DATA.W.SafetyStop
   //       R     #USER_DATA.W.FlyChange
   //       R     #USER_DATA.W.BrakeRelease
   //       R     #USER_DATA.W.ResetCount
   //       R     #USER_DATA.W.PresetRq
   //       R     #USER_DATA.W.HomeSearch
   //       R     #USER_DATA.W.ReverseHoming
   //       R     #USER_DATA.W.ReferenceCam
   //       R     #USER_DATA.W.ReferenceZero
   //       R     #USER_DATA.W.MDI_Continue
   //       R     #USER_DATA.W.SwLimitsEnable
   //       R     #USER_DATA.W.HwLimitsEnable
   //       R     #Run
   //       R     #Reverse
   //       R     #Positioning
   // 
   //       L     L#0
   //       T     #Speed
   //       T     #USER_DATA.W.Override
   //       T     #USER_DATA.W.Target
   //       T     #USER_DATA.W.Preset
   //       T     #USER_DATA.W.Acc
   //       T     #USER_DATA.W.Dec
   Rest: NOP   0;
   //    SET
   //    R     #IN_xDrive_EN
   //    R     #IN_xResetFaults
END_REGION

REGION Network 66 (STL): Restore AR1 & AR2 value
   //    L     #TMP_dOldValue_AR1
   //    LAR1
   //    L     #TMP_dOldValue_AR2
   //    LAR2
END_REGION
END_FUNCTION_BLOCK

FUNCTION_BLOCK "SINAMICS_SimpleDrive"   // FB53, LAD
TITLE = Sinamics drive manager
{ S7_Optimized_Access := 'FALSE' }
AUTHOR : Armitano
VERSION : 1.4
// Return value:
// * 0: OK
// Blocking message:
// * group 1 to 9: general error
// * group 10 to 19: system data error
//   * 10: Sinamics input/output addresses wrong or not setted
//   * 11: Maximum speed in Rpm wrong or not setted
//   * 12: Conversion coefficent for Rpm/mmMin wrong or not setted
//   * 13: Conversion coefficent for mmMin/Rpm wrong or not setted
//   * 14: Maximum acceleration wrong or not setted
//   * 15: Maximum deceleration wrong or not setted
//   * 19: Comunication telegram numxer unknown
// Warning message:
// * group 20 to 29: user data error
//   * 20: Reference cam signal + reference zero signal no possible
//   * 21: Run command + reverse command no possible
//   * 22: Preset speed at zero during run/reverse command
//   * 23: Run/reverse command during homing command no possible
//   * 24: Absolute positioining no possible without axes referenced
//   * 25: Preset override at zero during run/reverse command
// Other:
// * group 30 to 32: preset data error
//   * 30: Error during send preset value (Check parameters in Sys_Data)
//   * 31: Error during preset command (Check parameters in Sys_Data)
//   * 32: Error during saving preset command (Check Sys_Data)
//   * 34: Error during send preset homing (Check parameters in Sys_Data)
// * group 8000 to 9000: SFC20 code (Read the SFC20 Help)
   VAR_INPUT
      IN_xDrive_EN : Bool;   // Drive enable
      IN_xRun : Bool;   // Run forward
      IN_xReverse : Bool;   // Run backward
      IN_xRemoteRef : Bool;   // Remote reference
      IN_xResetFaults : Bool;   // Reset faults
      IN_dSpeed_mm_min : DInt;   // Speed reference [mm/min]
   END_VAR
   VAR_OUTPUT
      OUT_xFeedback : Bool;   // Feedback active
      OUT_xFaultPresent : Bool;   // Fault present
      OUT_iFaultCode : Int;   // Fault code
      OUT_iRetVal : Int;   // Return value in case of wrong configuration
   END_VAR
   VAR
      STC_tUSER_DATA : Struct   // User data (Extended functions commands for execute the application desired)
         tR : Struct
            xReadyfForSwitchOn : Bool;   // Ready for switch on
            xReadyToMove : Bool;   // Ready to move
            x2 : Bool;
            x3 : Bool;
            xAlarmPresent : Bool;   // Alarm present
            iAlarmCode : Int;   // Alarm code
            D6 : DInt;
            dActualSpeed_mm_min : DInt;   // Actual speed value [mm/min]
         END_STRUCT;
         tW : Struct
            xSafetyStop : Bool;   // Safety stop (OFF3)
            x1 : Bool;
            x2 : Bool;
            x3 : Bool;
            x4 : Bool;
            xBrakeRelease : Bool;   // Brake release
            x6 : Bool;
            x7 : Bool;
            x8 : Bool;
            x9 : Bool;
            x10 : Bool;
            x11 : Bool;
            x12 : Bool;
            x13 : Bool;
            x14 : Bool;
            x15 : Bool;
            i16 : Int := 100;
            d17 : DInt;
            d18 : DInt;
            rAcc_s : Real;   // Acceleration [s]
            rDec_s : Real;   // Deceleration [s]
         END_STRUCT;
      END_STRUCT;
      STC_tSYS_DATA : Struct   // System data (Info about applications type and HW config.)
         iIOAddress_MM : Int := -1;   // Input/Output addresses for motor module
         i2 : Int;
         i3 : Int;
         i4 : Int;
         i5 : Int;
         i6 : Int;
         i7 : Int;
         dMaxSpeed_rpm : DInt;   // MaxSpeed [rpm]
         d9 : DInt;
         d10 : DInt := L#1;
         d11 : DInt;
         d12 : DInt;
         d13 : DInt;
         rK_rpm_mmMin : Real;   // K Conversion from rpm to mm/min
         rK_mmMin_Rpm : Real;   // K Conversion from mm/min to rpm
         rMaxAcc_s : Real;   // MaxAcc [s]
         rMaxDec_s : Real;   // MaxDec [s]
         r18 : Real;
         r19 : Real;
      END_STRUCT;
      STC_tST : Struct
         x0 : Bool;
         x1 : Bool;
         x2 : Bool;
         x3 : Bool;
         x4 : Bool;
         x5 : Bool;
         x6 : Bool;
         x7 : Bool;
         x8 : Bool;
         x9 : Bool;
         x10 : Bool;
         x11 : Bool;
         x12 : Bool;
         x13 : Bool;
         x14 : Bool;
         x15 : Bool;
      END_STRUCT;
      STC_tOS_PN : Struct
         x0 : Bool;
         x1 : Bool;
         x2 : Bool;
         x3 : Bool;
         x4 : Bool;
         x5 : Bool;
         x6 : Bool;
         x7 : Bool;
         x8 : Bool;
         x9 : Bool;
         x10 : Bool;
         x11 : Bool;
         x12 : Bool;
         x13 : Bool;
         x14 : Bool;
         x15 : Bool;
      END_STRUCT;
      STC_tOS : Struct
         x0 : Bool;
         x1 : Bool;
         x2 : Bool;
         x3 : Bool;
         x4 : Bool;
         x5 : Bool;
         x6 : Bool;
         x7 : Bool;
         x8 : Bool;
         x9 : Bool;
         x10 : Bool;
         x11 : Bool;
         x12 : Bool;
         x13 : Bool;
         x14 : Bool;
         x15 : Bool;
      END_STRUCT;
      STC_tPH : Struct
         x0 : Bool;
         x1 : Bool;
         x2 : Bool;
         x3 : Bool;
         x4 : Bool;
         x5 : Bool;
         x6 : Bool;
         x7 : Bool;
         x8 : Bool;
         x9 : Bool;
         x10 : Bool;
         x11 : Bool;
         x12 : Bool;
         x13 : Bool;
         x14 : Bool;
         x15 : Bool;
      END_STRUCT;
      STC_tPROP : Struct
         i0 : Int;   // Previous cycle [ms]
         i1 : Int;
         i2 : Int;
         d3 : DInt;
         d4 : DInt;
         r5 : Real;
         r6 : Real;
         i7 : Int;
         i8 : Int;
         i9 : Int;
         i10 : Int;
         i11 : Int;
         d12 : DInt;
         d13 : DInt;
         r14 : Real;
         r15 : Real;
         i16 : Int;
         i17 : Int;